screen "IGG Digital Inputs" 1280x800, template "Template"
   on GenerateScreen: "TitleUpdater"()
   Button "HmiScreenItemData_1" at 1,1 size 150x43; TextOn 'Back'; TextOff 'Commissioning'
      on Release: ActivateScreen("Commissioning Main Page", 0)
   AlarmView "Alarm view_1" at 0,777 size 1280x23
   TextField "Text field_1" at 315,140 size 55x22; Text 'I0.0'
   TextField "Text field_2" at 315,176 size 55x22; Text 'I0.1'
   TextField "Text field_3" at 315,212 size 55x22; Text 'I0.2'
   TextField "Text field_4" at 315,248 size 55x22; Text 'I0.3'
   TextField "Text field_5" at 315,283 size 55x22; Text 'I0.4'
   TextField "Text field_6" at 315,319 size 55x22; Text 'I0.5'
   TextField "Text field_7" at 315,355 size 55x22; Text 'I0.6'
   TextField "Text field_8" at 315,391 size 55x22; Text 'I0.7'
   Circle "Circle_1" at 375,140 size 20x20
      Appearance <- "10_DI_Data_IGG_ESTOP_OK"
   Circle "Circle_2" at 375,176 size 20x20
      Appearance <- "10_DI_Data_E139_READY"
   Circle "Circle_3" at 375,212 size 20x20
      Appearance <- "10_DI_Data_E500A_TRIPPED"
   Circle "Circle_4" at 375,248 size 20x20
      Appearance <- "10_DI_Data_E500B_TRIPPED(1)"
   Circle "Circle_5" at 375,283 size 20x20
      Appearance <- "10_DI_Data_E500A_ENBLD(1)"
   Circle "Circle_6" at 375,319 size 20x20
      Appearance <- "10_DI_Data_E500B_ENBLD(1)"
   Circle "Circle_7" at 375,355 size 20x20
      Appearance <- "10_DI_Data_CV401_OPN"
   Circle "Circle_8" at 375,391 size 20x20
      Appearance <- "10_DI_Data_CV401_CLSD"
   TextField "Text field_9" at 332,108 size 49x26; Text 'I0'
   TextField "Text field_10" at 315,461 size 55x22; Text 'I1.0'
   TextField "Text field_11" at 315,497 size 55x22; Text 'I1.1'
   TextField "Text field_12" at 315,533 size 55x22; Text 'I1.2'
   TextField "Text field_13" at 315,569 size 55x22; Text 'I1.3'
   TextField "Text field_14" at 315,604 size 55x22; Text 'I1.4'
   TextField "Text field_15" at 315,640 size 55x22; Text 'I1.5'
   TextField "Text field_16" at 315,676 size 55x22; Text 'I1.6'
   TextField "Text field_17" at 315,712 size 55x22; Text 'I1.7'
   Circle "Circle_9" at 375,461 size 20x20
      Appearance <- "10_DI_Data_CV321_OPN"
   Circle "Circle_10" at 375,497 size 20x20
      Appearance <- "10_DI_Data_CV321_CLSD"
   Circle "Circle_11" at 375,533 size 20x20
      Appearance <- "10_DI_Data_CV322_OPN"
   Circle "Circle_12" at 375,569 size 20x20
      Appearance <- "10_DI_Data_CV322_CLSD"
   Circle "Circle_13" at 375,604 size 20x20
      Appearance <- "10_DI_Data_CV311_OPN"
   Circle "Circle_14" at 375,640 size 20x20
      Appearance <- "10_DI_Data_CV311_CLSD"
   Circle "Circle_15" at 375,676 size 20x20
      Appearance <- "10_DI_Data_CV312_OPN"
   Circle "Circle_16" at 375,712 size 20x20
      Appearance <- "10_DI_Data_CV312_CLSD"
   TextField "Text field_18" at 332,429 size 49x26; Text 'I1'
   TextField "Text field_19" at 657,141 size 55x22; Text 'I2.0'
   TextField "Text field_20" at 657,177 size 55x22; Text 'I2.1'
   TextField "Text field_21" at 657,213 size 55x22; Text 'I2.2'
   TextField "Text field_22" at 657,249 size 55x22; Text 'I2.3'
   TextField "Text field_23" at 657,284 size 55x22; Text 'I2.4'
   TextField "Text field_24" at 657,320 size 55x22; Text 'I2.5'
   TextField "Text field_25" at 657,356 size 55x22; Text 'I2.6'
   TextField "Text field_26" at 657,392 size 55x22; Text 'I2.7'
   Circle "Circle_17" at 717,141 size 20x20
      Appearance <- "10_DI_Data_BC_PLC_PWR_OK"
   Circle "Circle_18" at 717,177 size 20x20
      Appearance <- "10_DI_Data_IGG_VNT_PWR_OK"
   Circle "Circle_19" at 717,213 size 20x20
      Appearance <- "10_DI_Data_MCC_VNT_PWR_OK"
   Circle "Circle_20" at 717,249 size 20x20
      Appearance <- "10_DI_Data_7T1_PWR_OK"
   Circle "Circle_21" at 717,284 size 20x20
      Appearance <- "10_DI_Data_7T2_PWR_OK"
   Circle "Circle_22" at 717,320 size 20x20
      Appearance <- "10_DI_Data_7T3_PWR_OK"
   Circle "Circle_23" at 717,356 size 20x20
      Appearance <- "10_DI_Data_MAINTD_24VDC_PWR_OK"
   Circle "Circle_24" at 717,392 size 20x20
      Appearance <- "10_DI_Data_SFTY_SYS_IL"
   TextField "Text field_27" at 674,109 size 49x26; Text 'I2'
   TextField "Text field_37" at 315,66 size 254x26; Text 'IGG System PLC (Rack 1)'
   TextField "Text field_28" at 657,459 size 55x22; Text 'I3.0'
   TextField "Text field_29" at 657,495 size 55x22; Text 'I3.1'
   TextField "Text field_30" at 657,531 size 55x22; Text 'I3.2'
   TextField "Text field_31" at 657,567 size 55x22; Text 'I3.3'
   TextField "Text field_32" at 657,602 size 55x22; Text 'I3.4'
   TextField "Text field_33" at 657,638 size 55x22; Text 'I3.5'
   TextField "Text field_34" at 657,674 size 55x22; Text 'I3.6'
   TextField "Text field_35" at 657,710 size 55x22; Text 'I3.7'
   Circle "Circle_25" at 717,459 size 20x20
      Appearance <- "10_DI_Data_CV432_OPN"
   Circle "Circle_26" at 717,495 size 20x20
      Appearance <- "10_DI_Data_CV432_CLSD"
   Circle "Circle_27" at 717,531 size 20x20
      Appearance <- "10_DI_Data_CV431_OPN"
   Circle "Circle_28" at 717,567 size 20x20
      Appearance <- "10_DI_Data_CV431_CLSD"
   Circle "Circle_29" at 717,602 size 20x20
      Appearance <- "10_DI_Data_E139_RUNNING(1)"
   Circle "Circle_30" at 717,638 size 20x20
      Appearance <- "10_DI_Data_E139_VSD_FLT"
   Circle "Circle_31" at 717,674 size 20x20
      Appearance <- "10_DI_Data_MCCP_5PG1_OK"
   Circle "Circle_32" at 717,710 size 20x20
      Appearance <- "10_DI_Data_R1_SPR_DI_3_7"
   TextField "Text field_36" at 674,427 size 49x26; Text 'I3'
   TextField "Text field_75" at 408,140 size 200x22; Text 'IGG E-Stop Healthy'
   TextField "Text field_76" at 408,175 size 200x22; Text 'CA Blower Ready E139'
   TextField "Text field_77" at 408,211 size 200x22; Text 'Fuel Pump 1 Tripped E500A'
   TextField "Text field_78" at 408,247 size 200x22; Text 'Fuel Pump 2 Tripped E500B'
   TextField "Text field_79" at 408,283 size 200x22; Text 'Fuel Pump 1 Enabled E500A'
   TextField "Text field_80" at 408,319 size 200x22; Text 'Fuel Pump 2 Enabled E500B'
   TextField "Text field_81" at 408,355 size 200x22; Text 'IG Supply Valve Open CV401'
   TextField "Text field_82" at 408,391 size 200x22; Text 'IG Supply Valve Closed CV401'
   TextField "Text field_83" at 408,460 size 200x22; Text 'DTB Valve Open CV321'
   TextField "Text field_84" at 408,496 size 200x22; Text 'DTB Valve Closed CV321'
   TextField "Text field_85" at 408,532 size 200x22; Text 'CSW Drain Valve Open CV322'
   TextField "Text field_86" at 408,568 size 200x22; Text 'CSW Drain Valve Closed CV322'
   TextField "Text field_87" at 408,604 size 200x22; Text 'CSW Valve Open CV311'
   TextField "Text field_88" at 408,640 size 200x22; Text 'CSW Valve Closed CV311'
   TextField "Text field_89" at 408,676 size 200x22; Text 'Flue Gas S CSW Valve Open CV312'
   TextField "Text field_90" at 408,712 size 200x22; Text 'Flue Gas S CSW Valve Closed CV312'
   TextField "Text field_91" at 748,139 size 200x22; Text 'BC PLC Power Healthy'
   TextField "Text field_92" at 748,175 size 200x22; Text 'IGG Vent Power Healthy'
   TextField "Text field_93" at 748,211 size 200x22; Text 'MCC Vent Power Healthy'
   TextField "Text field_94" at 748,247 size 200x22; Text '7T1 Power Healthy'
   TextField "Text field_95" at 748,283 size 200x22; Text '7T2 Power Healthy'
   TextField "Text field_96" at 748,319 size 200x22; Text '7T3 Power Healthy'
   TextField "Text field_97" at 748,355 size 200x22; Text 'Maintained 24V Power'
   TextField "Text field_98" at 748,392 size 200x22; Text 'Safety System Interlock'
   TextField "Text field_99" at 749,458 size 200x22; Text 'CB IG Supply Valve Open CV432'
   TextField "Text field_100" at 749,494 size 200x22; Text 'CB IG Supply Valve Closed CV432'
   TextField "Text field_101" at 749,530 size 200x22; Text 'BWTS IG Supply Open CV431'
   TextField "Text field_102" at 749,566 size 200x22; Text 'BWTS IG Supply Closed CV431'
   TextField "Text field_103" at 749,602 size 200x22; Text 'CA Blower Running E139'
   TextField "Text field_104" at 749,638 size 200x22; Text 'VSD Fault'
   TextField "Text field_105" at 749,674 size 200x22; Text 'Correct Phase Rotation'
   TextField "Text field_106" at 749,711 size 200x22; Text 'Spare Input'
   Group "Group" at 750,42 size 373x50
   Button "HmiScreenItemData_8" at 764,46 size 355x40; TextOn 'Back'; TextOff 'Text'
   TextField "Screen title" at 750,42 size 373x50; Text 'Screen title'

screen "BC Digital Outputs" 1280x800, template "Template"
   on GenerateScreen: "TitleUpdater"()
   Button "HmiScreenItemData_1" at 1,1 size 150x43; TextOn 'Back'; TextOff 'Commissioning'
      on Release: ActivateScreen("Commissioning Main Page", 0)
   AlarmView "Alarm view_1" at 0,777 size 1280x23
   TextField "Text field_37" at 319,170 size 287x26; Text 'Burner Control PLC (Rack 2)'
   TextField "Text field_38" at 384,239 size 55x22; Text 'Q0.0'
   TextField "Text field_39" at 384,290 size 55x22; Text 'Q0.1'
   TextField "Text field_40" at 384,342 size 55x22; Text 'Q0.2'
   TextField "Text field_41" at 384,394 size 55x22; Text 'Q0.3'
   TextField "Text field_42" at 384,446 size 55x22; Text 'Q0.4'
   TextField "Text field_43" at 384,498 size 55x22; Text 'Q0.5'
   TextField "Text field_44" at 384,550 size 55x22; Text 'Q0.6'
   TextField "Text field_45" at 384,602 size 55x22; Text 'Q0.7'
   Circle "Circle_33" at 443,239 size 20x20
      Appearance <- "14_DQ_Data_200CV127ControlOut"
   Circle "Circle_34" at 443,290 size 20x20
      Appearance <- "14_DQ_Data_200CV124ControlOut"
   Circle "Circle_35" at 443,342 size 20x20
      Appearance <- "14_DQ_Data_200CV215ControlOut"
   Circle "Circle_36" at 443,394 size 20x20
      Appearance <- "14_DQ_Data_200CV216ControlOut"
   Circle "Circle_37" at 443,446 size 20x20
      Appearance <- "14_DQ_Data_200CV114ControlOut"
   Circle "Circle_38" at 443,498 size 20x20
      Appearance <- "14_DQ_Data_200CV206ControlOut"
   Circle "Circle_39" at 443,550 size 20x20
      Appearance <- "14_DQ_Data_200CV207ControlOut"
   Circle "Circle_40" at 443,602 size 20x20
      Appearance <- "14_DQ_Data_E131ControlOut"
   TextField "Text field_46" at 398,206 size 49x26; Text 'Q0'
   TextField "Text field_47" at 703,239 size 55x22; Text 'Q1.0'
   TextField "Text field_48" at 703,290 size 55x22; Text 'Q1.1'
   TextField "Text field_49" at 703,342 size 55x22; Text 'Q1.2'
   TextField "Text field_50" at 703,394 size 55x22; Text 'Q1.3'
   TextField "Text field_51" at 703,446 size 55x22; Text 'Q1.4'
   TextField "Text field_52" at 703,498 size 55x22; Text 'Q1.5'
   TextField "Text field_53" at 703,550 size 55x22; Text 'Q1.6'
   TextField "Text field_54" at 703,602 size 55x22; Text 'Q1.7'
   Circle "Circle_41" at 763,239 size 20x20
      Appearance <- "51_SLAVE_STATUS_P301_ENBLD"
   Circle "Circle_42" at 763,290 size 20x20
      Appearance <- "14_DQ_Data_X001ControlOut"
   Circle "Circle_43" at 763,341 size 20x20
      Appearance <- "14_DQ_Data_R2_SPR_DQ_1_2"
   Circle "Circle_44" at 763,394 size 20x20
      Appearance <- "14_DQ_Data_R2_SPR_DQ_1_3"
   Circle "Circle_45" at 763,446 size 20x20
      Appearance <- "14_DQ_Data_R2_SPR_DQ_1_4"
   Circle "Circle_46" at 763,500 size 20x20
      Appearance <- "14_DQ_Data_R2_SPR_DQ_1_5"
   Circle "Circle_47" at 763,551 size 20x20
      Appearance <- "14_DQ_Data_R2_SPR_DQ_1_6"
   Circle "Circle_48" at 763,602 size 20x20
      Appearance <- "14_DQ_Data_P305ControlOut"
   TextField "Text field_55" at 716,206 size 49x26; Text 'Q1'
   Button "Button_1" at 321,231 size 60x35; TextOff 'Override'
      on Press: InvertBit("80_From_HMI_MAN_DQ_0_0(1)")
      Visibility <- "82_To_HMI_CRNT_MODE_IGG"
   Button "Button_2" at 321,283 size 60x35; TextOff 'Override'
      on Press: InvertBit("80_From_HMI_MAN_DQ_0_1(1)")
      Visibility <- "82_To_HMI_CRNT_MODE_IGG"
   Button "Button_3" at 321,335 size 60x35; TextOff 'Override'
      on Press: InvertBit("80_From_HMI_MAN_DQ_0_2(1)")
      Visibility <- "82_To_HMI_CRNT_MODE_IGG"
   Button "Button_4" at 321,387 size 60x35; TextOff 'Override'
      on Press: InvertBit("80_From_HMI_MAN_DQ_0_3(1)")
      Visibility <- "82_To_HMI_CRNT_MODE_IGG"
   Button "Button_5" at 321,439 size 60x35; TextOff 'Override'
      on Press: InvertBit("80_From_HMI_MAN_DQ_0_4(1)")
      Visibility <- "82_To_HMI_CRNT_MODE_IGG"
   Button "Button_6" at 321,491 size 60x35; TextOff 'Override'
      on Press: InvertBit("80_From_HMI_MAN_DQ_0_5(1)")
      Visibility <- "82_To_HMI_CRNT_MODE_IGG"
   Button "Button_7" at 321,543 size 60x35; TextOff 'Override'
      on Press: InvertBit("80_From_HMI_MAN_DQ_0_6(1)")
      Visibility <- "82_To_HMI_CRNT_MODE_IGG"
   Button "Button_8" at 639,283 size 60x35; TextOff 'Override'
      on Press: InvertBit("80_From_HMI_MAN_DQ_1_1(1)")
      Visibility <- "82_To_HMI_CRNT_MODE_IGG"
   Button "Button_13" at 321,596 size 60x35; TextOff 'Override'
      on Press: InvertBit("80_From_HMI_MAN_DQ_0_7")
      Visibility <- "82_To_HMI_CRNT_MODE_IGG"
   TextField "Text field_72" at 465,239 size 170x22; Text 'Test Pressure Valve CV127'
   TextField "Text field_73" at 465,290 size 170x22; Text 'Pilot B Ign Valve CV124'
   TextField "Text field_75" at 465,342 size 170x22; Text 'Pilot B Fuel Valve 1 CV215'
   TextField "Text field_76" at 465,394 size 170x22; Text 'Pilot B Fuel Valve 2 CV215'
   TextField "Text field_77" at 465,446 size 170x22; Text 'Main B Atom Air Vlv CV114'
   TextField "Text field_78" at 465,498 size 170x22; Text 'Main B Fuel Valve 1 CV205'
   TextField "Text field_79" at 465,550 size 170x22; Text 'Main B Fuel Valve 2 CV206'
   TextField "Text field_80" at 465,602 size 170x22; Text 'IA Comp E131'
   TextField "Text field_81" at 792,238 size 170x22; Text 'CSW Pump P301'
   TextField "Text field_82" at 792,290 size 170x22; Text 'Ignitor X001'
   TextField "Text field_86" at 792,342 size 170x22; Text 'Spare Output'
   TextField "Text field_87" at 792,394 size 170x22; Text 'Spare Output'
   TextField "Text field_88" at 792,446 size 170x22; Text 'Spare Output'
   TextField "Text field_89" at 792,498 size 170x22; Text 'Spare Output'
   TextField "Text field_90" at 792,550 size 170x22; Text 'Spare Output'
   TextField "Text field_91" at 792,602 size 170x22; Text 'Fresh Water Pump'
   Button "Button_26" at 639,231 size 60x35; TextOff 'Override'
      on Press: InvertBit("80_From_HMI_MAN_DQ_1_0")
      Visibility <- "82_To_HMI_CRNT_MODE_IGG"
   Button "Button_27" at 639,335 size 60x35; TextOff 'Override'
      on Press: InvertBit("80_From_HMI_MAN_DQ_1_2(1)")
      Visibility <- "82_To_HMI_CRNT_MODE_IGG"
   Button "Button_28" at 639,439 size 60x35; TextOff 'Override'
      on Press: InvertBit("80_From_HMI_MAN_DQ_1_4(1)")
      Visibility <- "82_To_HMI_CRNT_MODE_IGG"
   Button "Button_29" at 639,387 size 60x35; TextOff 'Override'
      on Press: InvertBit("80_From_HMI_MAN_DQ_1_3(1)")
      Visibility <- "82_To_HMI_CRNT_MODE_IGG"
   Button "Button_30" at 639,491 size 60x35; TextOff 'Override'
      on Press: InvertBit("80_From_HMI_MAN_DQ_1_5(1)")
      Visibility <- "82_To_HMI_CRNT_MODE_IGG"
   Button "Button_31" at 639,543 size 60x35; TextOff 'Override'
      on Press: InvertBit("80_From_HMI_MAN_DQ_1_6")
      Visibility <- "82_To_HMI_CRNT_MODE_IGG"
   Button "Button_32" at 639,596 size 60x35; TextOff 'Override'
      on Press: InvertBit("80_From_HMI_MAN_DQ_1_7(1)")
      Visibility <- "82_To_HMI_CRNT_MODE_IGG"
   Group "Group" at 455,41 size 373x50
   Button "HmiScreenItemData_8" at 469,45 size 355x40; TextOn 'Back'; TextOff 'Text'
   TextField "Screen title" at 455,41 size 373x50; Text 'Screen title'

screen "BC Analogue Inputs" 1280x800, template "Template"
   on GenerateScreen: "TitleUpdater"()
   Button "HmiScreenItemData_1" at 1,1 size 150x43; TextOn 'Back'; TextOff 'Commissioning'
      on Release: ActivateScreen("Commissioning Main Page", 0)
   Button "Button_1" at 34,732 size 100x35; TextOn 'BWTS Digital Inputs'; TextOff 'Back'
      on Click: ActivateScreen("IGG Analogue Inputs", 0)
   TextField "Text field_39" at 34,688 size 171x62; Text 'To IGG Analogue Inputs'
   AlarmView "Alarm view_1" at 0,777 size 1280x23
   Group "Group_1" at 455,41 size 373x50
   TextField "Text field_26" at 607,234 size 64x20; Text 'Reading'
   TextField "Text field_27" at 680,234 size 68x20; Text 'Low Low'
   TextField "Text field_28" at 761,234 size 37x20; Text 'Low'
   TextField "Text field_29" at 829,234 size 37x20; Text 'High'
   TextField "Text field_30" at 879,234 size 74x20; Text 'High High'
   TextField "Text field_31" at 755,211 size 76x20; Text 'Setpoints'
   TextField "Text field_42" at 450,234 size 89x20; Text 'Description'
   TextField "Text field_44" at 340,234 size 37x20; Text 'AI'
   TextField "Text field_53" at 335,202 size 364x26; Text 'Burner Control System PLC (Rack 2)'
   TextField "Text field_35" at 381,576 size 220x22; Text 'E-700 - Inert Gas Soot Content'
   IOField "I/O field_61" at 608,576 size 70x22; FormatPattern 999.99; Unit  %
      ProcessValue <- "12_AI_Data_E700SootContentIn"
   IOField "I/O field_62" at 682,576 size 60x22; FormatPattern 9.9
   TextField "Text field_36" at 328,576 size 50x22; Text 'IW110'
   IOField "I/O field_64" at 750,576 size 60x22; Authorization "Parameter Change"; FormatPattern 99.9
      ProcessValue <- "84_Setpoints_TX700_Low"
   IOField "I/O field_65" at 818,576 size 60x22; Authorization "Parameter Change"; FormatPattern 99.9
      ProcessValue <- "84_Setpoints_TX700_High"
   IOField "I/O field_63" at 886,576 size 60x22; FormatPattern 9.9
   TextField "Text field_1" at 381,536 size 220x22; Text 'E-600 CB - Oxygen Analyser Content'
   IOField "I/O field_2" at 750,536 size 60x22; Authorization "Parameter Change"; FormatPattern 9.99
      ProcessValue <- "84_Setpoints_E600_CB_Low"
   TextField "Text field_2" at 328,536 size 50x22; Text 'IW108'
   IOField "I/O field_8" at 818,536 size 60x22; Authorization "Parameter Change"; FormatPattern 9.99
      ProcessValue <- "84_Setpoints_E600_CB_High"
   IOField "I/O field_1" at 682,536 size 60x22; Authorization "Parameter Change"; FormatPattern 9.99
      ProcessValue <- "84_Setpoints_E600_CB_LowLow"
   IOField "I/O field_9" at 886,536 size 60x22; Authorization "Parameter Change"; FormatPattern 9.99
      ProcessValue <- "84_Setpoints_E600_CB_HighHigh"
   TextField "Text field_33" at 381,496 size 220x22; Text 'E-600 BWTS - Oxygen Analyser Content'
   IOField "I/O field_56" at 608,496 size 70x22; FormatPattern 99.99; Unit  %
      ProcessValue <- "12_AI_Data_E600O2ContentIn"
   IOField "I/O field_58" at 750,496 size 60x22; Authorization "Parameter Change"; FormatPattern 9.99
      ProcessValue <- "84_Setpoints_E600_BWT_Low"
   TextField "Text field_34" at 328,496 size 50x22; Text 'IW108'
   IOField "I/O field_59" at 818,496 size 60x22; Authorization "Parameter Change"; FormatPattern 9.99
      ProcessValue <- "84_Setpoints_E600_BWT_High"
   IOField "I/O field_10" at 886,496 size 60x22; Authorization "Parameter Change"; FormatPattern 9.99
      ProcessValue <- "84_Setpoints_E600_BWT_HighHigh"
   IOField "I/O field_11" at 682,496 size 60x22; Authorization "Parameter Change"; FormatPattern 9.99
      ProcessValue <- "84_Setpoints_E600_BWT_LowLow"
   TextField "Text field_25" at 381,456 size 220x22; Text 'TIT-202 - Inlet Fuel Temperature'
   IOField "I/O field_51" at 608,456 size 70x22; FormatPattern s999.9; Unit  °C
      ProcessValue <- "12_AI_Data_TIT202In_SCALED"
   TextField "Text field_32" at 328,456 size 50x22; Text 'IW106'
   IOField "I/O field_52" at 682,456 size 60x22; Authorization "Parameter Change"; FormatPattern s999.9
      ProcessValue <- "84_Setpoints_TIT202_LowLow"
   IOField "I/O field_53" at 750,456 size 60x22; Authorization "Parameter Change"; FormatPattern s999.9
      ProcessValue <- "84_Setpoints_TIT202_Low"
   IOField "I/O field_54" at 818,456 size 60x22; Authorization "Parameter Change"; FormatPattern s999.9
      ProcessValue <- "84_Setpoints_TIT202_High"
   IOField "I/O field_55" at 886,456 size 60x22; Authorization "Parameter Change"; FormatPattern s999.9
      ProcessValue <- "84_Setpoints_TIT202_HighHigh"
   TextField "Text field_73" at 381,417 size 220x22; Text 'PIT-204 - IGG Inlet Fuel Pressure'
   IOField "I/O field_146" at 608,417 size 70x22; FormatPattern 99.9; Unit  Bar
      ProcessValue <- "12_AI_Data_PIT204In_SCALED"
   TextField "Text field_74" at 328,417 size 50x22; Text 'IW104'
   IOField "I/O field_147" at 682,417 size 60x22; Authorization "Parameter Change"; FormatPattern 99.9
      ProcessValue <- "84_Setpoints_PIT204_LowLow(2)"
   IOField "I/O field_148" at 750,417 size 60x22; Authorization "Parameter Change"; FormatPattern 99.9
      ProcessValue <- "84_Setpoints_PIT204_Low(2)"
   IOField "I/O field_149" at 818,417 size 60x22; Authorization "Parameter Change"; FormatPattern 99.9
      ProcessValue <- "84_Setpoints_PIT204_High(2)"
   IOField "I/O field_150" at 886,417 size 60x22; Authorization "Parameter Change"; FormatPattern 99.9
      ProcessValue <- "84_Setpoints_PIT204_HighHigh(2)"
   TextField "Text field_71" at 381,378 size 220x22; Text 'PIT-112 - Inlet IA Compressor Pressure'
   TextField "Text field_72" at 328,378 size 50x22; Text 'IW102'
   IOField "I/O field_3" at 608,378 size 70x22; FormatPattern 99.9; Unit  Bar
      ProcessValue <- "12_AI_Data_PIT112In_SCALED"
   IOField "I/O field_4" at 682,378 size 60x22; Authorization "Parameter Change"; FormatPattern 99.9
      ProcessValue <- "84_Setpoints_PIT112_LowLow"
   IOField "I/O field_5" at 750,378 size 60x22; Authorization "Parameter Change"; FormatPattern 99.9
      ProcessValue <- "84_Setpoints_PIT112_Low"
   IOField "I/O field_6" at 818,378 size 60x22; Authorization "Parameter Change"; FormatPattern 99.9
      ProcessValue <- "84_Setpoints_PIT112_High"
   IOField "I/O field_7" at 886,378 size 60x22; Authorization "Parameter Change"; FormatPattern 99.9
      ProcessValue <- "84_Setpoints_PIT112_HighHigh"
   TextField "Text field_69" at 381,338 size 220x22; Text 'PIT-113 - Main Atom. Air Pressure'
   IOField "I/O field_136" at 608,338 size 70x22; FormatPattern 99.9; Unit  Bar
      ProcessValue <- "12_AI_Data_PIT113In_SCALED"
   TextField "Text field_70" at 328,338 size 50x22; Text 'IW100'
   IOField "I/O field_137" at 682,338 size 60x22; Authorization "Parameter Change"; FormatPattern 99.9
      ProcessValue <- "84_Setpoints_PIT113_LowLow"
   IOField "I/O field_138" at 750,338 size 60x22; Authorization "Parameter Change"; FormatPattern 99.9
      ProcessValue <- "84_Setpoints_PIT113_Low"
   IOField "I/O field_139" at 818,338 size 60x22; Authorization "Parameter Change"; FormatPattern 99.9
      ProcessValue <- "84_Setpoints_PIT113_High"
   IOField "I/O field_140" at 886,338 size 60x22; Authorization "Parameter Change"; FormatPattern 99.9
      ProcessValue <- "84_Setpoints_PIT113_HighHigh"
   TextField "Text field_67" at 381,299 size 220x22; Text 'FD-001 - Flame Signal'
   IOField "I/O field_131" at 608,299 size 70x22; FormatPattern 999.9; Unit  %
      ProcessValue <- "12_AI_Data_FD001FlameSignalIn"
   IOField "I/O field_134" at 818,299 size 60x22; FormatPattern s99.9
   IOField "I/O field_135" at 886,299 size 60x22; FormatPattern s99.9
   TextField "Text field_68" at 328,299 size 50x22; Text 'IW98'
   IOField "I/O field_132" at 682,299 size 60x22; Authorization "Parameter Change"; FormatPattern 999.9
      ProcessValue <- "84_Setpoints_FD001_LowLow"
   IOField "I/O field_133" at 750,299 size 60x22; Authorization "Parameter Change"; FormatPattern 999.9
      ProcessValue <- "84_Setpoints_FD001_Low"
   TextField "Text field_65" at 381,260 size 220x22; Text 'PIT-205 - IGG Main Fuel Pressure'
   IOField "I/O field_126" at 608,260 size 70x22; FormatPattern 99.9; Unit  Bar
      ProcessValue <- "12_AI_Data_PIT205In_SCALED"
   TextField "Text field_66" at 328,260 size 50x22; Text 'IW96'
   IOField "I/O field_127" at 682,260 size 60x22; Authorization "Parameter Change"; FormatPattern 99.9
      ProcessValue <- "84_Setpoints_PIT205_LowLow"
   IOField "I/O field_128" at 750,260 size 60x22; Authorization "Parameter Change"; FormatPattern 99.9
      ProcessValue <- "84_Setpoints_PIT205_Low"
   IOField "I/O field_129" at 818,260 size 60x22; Authorization "Parameter Change"; FormatPattern 99.9
      ProcessValue <- "84_Setpoints_PIT205_High"
   IOField "I/O field_130" at 886,260 size 60x22; Authorization "Parameter Change"; FormatPattern 99.9
      ProcessValue <- "84_Setpoints_PIT205_HighHigh"
   Button "HmiScreenItemData_8" at 469,45 size 355x40; TextOn 'Back'; TextOff 'Text'
   TextField "Screen title" at 455,41 size 373x50; Text 'Screen title'

screen "IGG Analogue Outputs" 1280x800, template "Template"
   on GenerateScreen: "TitleUpdater"()
   Button "HmiScreenItemData_1" at 1,1 size 150x43; TextOn 'Back'; TextOff 'Commissioning'
      on Release: ActivateScreen("Commissioning Main Page", 0)
   Button "Button_15" at 34,732 size 100x35; TextOn 'BWTS Digital Inputs'; TextOff 'Back'
      on Click: ActivateScreen("BC Analogue Inputs", 0)
   AlarmView "Alarm view_1" at 0,777 size 1280x23
   TextField "Text field_82" at 481,361 size 220x22; Text 'Vent Valve Position Control'
   TextField "Text field_90" at 750,332 size 64x20; Text 'Reading'
   IOField "I/O field_2" at 749,363 size 70x22; FormatPattern 9999; Unit %
      ProcessValue <- "16_AQ_Data_CV403_CNTRL"
   TextField "Text field_6" at 428,361 size 53x22; Text 'QW98'
   TextField "Text field_7" at 480,438 size 220x22; Text 'Spare'
   TextField "Text field_41" at 553,332 size 89x20; Text 'Description'
   TextField "Text field_43" at 437,332 size 37x20; Text 'AO'
   TextField "Text field_52" at 437,299 size 333x26; Text 'IGG Control System PLC (Rack 1)'
   TextField "Text field_25" at 480,399 size 220x22; Text 'CA Blower Speed Control'
   IOField "I/O field_51" at 749,398 size 70x22; FormatPattern 9999; Unit RPM
      ProcessValue <- "16_AQ_Data_E139_SPEED"
   TextField "Text field_32" at 427,399 size 53x22; Text 'QW100'
   Button "Button_24" at 716,359 size 29x26; TextOff '+'
      Visibility <- "82_To_HMI_CRNT_MODE_IGG"
      on Press: function_b14e0dd5("80_From_HMI_MAN_AQ_INC_98(1)", 0)
   Button "Button_25" at 824,359 size 29x26; TextOff '-'
      Visibility <- "82_To_HMI_CRNT_MODE_IGG"
      on Press: function_b14e0dd5("80_From_HMI_MAN_AQ_DEC_98(1)", 0)
   Button "Button_1" at 717,397 size 29x26; TextOff '+'
      Visibility <- "82_To_HMI_CRNT_MODE_IGG"
      on Press: function_b14e0dd5("80_From_HMI_MAN_AQ_INC_100", 0)
   Button "Button_2" at 825,397 size 29x26; TextOff '-'
      Visibility <- "82_To_HMI_CRNT_MODE_IGG"
      on Press: function_b14e0dd5("80_From_HMI_MAN_AQ_DEC_100", 0)
   Button "Button_3" at 715,434 size 29x26; TextOff '+'
      on Click: SetBit("80_From_HMI_MAN_AQ_INC_102(1)")
      Visibility <- "82_To_HMI_CRNT_MODE_IGG"
   Button "Button_4" at 823,434 size 29x26; TextOff '-'
      on Click: SetBit("80_From_HMI_MAN_AQ_DEC_102(1)")
      Visibility <- "82_To_HMI_CRNT_MODE_IGG"
   Button "Button_5" at 716,475 size 29x26; TextOff '+'
      on Click: SetBit("80_From_HMI_MAN_AQ_INC_104")
      Visibility <- "82_To_HMI_CRNT_MODE_IGG"
   Button "Button_6" at 824,475 size 29x26; TextOff '-'
      on Click: SetBit("80_From_HMI_MAN_AQ_DEC_104")
      Visibility <- "82_To_HMI_CRNT_MODE_IGG"
   IOField "I/O field_1" at 749,438 size 70x22; FormatPattern 9.9; Unit  
      ProcessValue <- "16_AQ_Data_R1_SPR_AQ_102"
   IOField "I/O field_3" at 750,478 size 70x22; FormatPattern 9.9; Unit  
      ProcessValue <- "16_AQ_Data_R1_SPR_AQ_104"
   TextField "Text field_1" at 480,478 size 220x22; Text 'Spare'
   TextField "Text field_2" at 428,438 size 53x22; Text 'QW102'
   TextField "Text field_3" at 427,478 size 53x22; Text 'QW104'
   Group "Group" at 455,41 size 373x50
   Button "HmiScreenItemData_8" at 469,45 size 355x40; TextOn 'Back'; TextOff 'Text'
   TextField "Screen title" at 455,41 size 373x50; Text 'Screen title'

screen "IGG Target Setpoints" 1280x800, template "Template"
   on GenerateScreen: "TitleUpdater"()
   Button "HmiScreenItemData_1" at 1,1 size 150x43; TextOn 'Back'; TextOff 'Commissioning'
      on Release: ActivateScreen("Commissioning Main Page", 0)
   AlarmView "Alarm view_1" at 0,777 size 1280x23
   TextField "Text field_25" at 394,430 size 407x22; Text 'PIT-113: IGG Main Atom Air Pressure Target'
   TextField "Text field_29" at 814,210 size 68x20; Text 'Setpoint'
   TextField "Text field_33" at 393,468 size 408x22; Text 'PIT-205: IGG Main Fuel Pressure Target'
   IOField "I/O field_58" at 816,468 size 60x22; Authorization "Parameter Change"; FormatPattern 999.99
      ProcessValue <- "84_Setpoints_PIT205_Target(1)"
   TextField "Text field_35" at 394,552 size 406x22; Text 'E-600: O2 Cargo Blanketing Target'
   TextField "Text field_65" at 394,236 size 411x22; Text 'PIT-402: IG Outlet Pressure Pilot Target'
   TextField "Text field_67" at 394,274 size 410x22; Text 'PIT-402: IG Outlet Pressure Main Target'
   TextField "Text field_69" at 395,313 size 407x22; Text 'PIT-402: IG Outlet Pressure Post Target Start'
   TextField "Text field_71" at 395,352 size 406x22; Text 'PIT-402: IG Outlet Pressure Post Target Maximum'
   TextField "Text field_73" at 395,391 size 407x22; Text 'FD-001: Igniter Target'
   TextField "Text field_42" at 394,210 size 89x20; Text 'Description'
   IOField "I/O field_128" at 816,236 size 60x22; Authorization "Parameter Change"; FormatPattern 999.9
      ProcessValue <- "84_Setpoints_PIT402_Pilot_Target(1)"
   IOField "I/O field_133" at 816,274 size 60x22; Authorization "Parameter Change"; FormatPattern 999.9
      ProcessValue <- "84_Setpoints_PIT402_Main_Target(1)"
   IOField "I/O field_138" at 816,313 size 60x22; Authorization "Parameter Change"; FormatPattern 999.9
      ProcessValue <- "84_Setpoints_PIT402_Post_Target_Start"
   IOField "I/O field_53" at 816,430 size 60x22; Authorization "Parameter Change"; FormatPattern 999.9
      ProcessValue <- "84_Setpoints_PIT113_Pilot_Target(1)"
   IOField "I/O field_148" at 816,391 size 60x22; Authorization "Parameter Change"; FormatPattern 999.9
      ProcessValue <- "84_Setpoints_FD001_Min"
   IOField "I/O field_64" at 816,552 size 60x22; Authorization "Parameter Change"; FormatPattern 99.9
      ProcessValue <- "84_Setpoints_E600_CB_Target"
   TextField "Text field_53" at 393,184 size 213x26; Text 'IGG Target Setpoints'
   IOField "I/O field_5" at 815,352 size 60x22; Authorization "Parameter Change"; FormatPattern 999.9
      ProcessValue <- "84_Setpoints_PIT401_Post_Target_Max"
   TextField "Text field_1" at 394,510 size 406x22; Text 'E-600: O2 Ballast Water Treatment Target'
   IOField "I/O field_2" at 816,510 size 60x22; Authorization "Parameter Change"; FormatPattern 9.99
      ProcessValue <- "84_Setpoints_E600_BWT_Target"
   TextField "Text field_2" at 394,595 size 406x22; Text 'PIT-402 Target Ramp Time (s)'
   IOField "I/O field_1" at 816,595 size 60x22; Authorization "Parameter Change"; FormatPattern 999
      ProcessValue <- "86_Times_PIT402_Ramp_Seconds"
   Group "Group" at 455,41 size 373x50
   Button "HmiScreenItemData_8" at 469,45 size 355x40; TextOn 'Back'; TextOff 'Text'
   TextField "Screen title" at 455,41 size 373x50; Text 'Screen title'

screen "IGG Process Times" 1280x800, template "Template"
   on GenerateScreen: "TitleUpdater"()
   Button "HmiScreenItemData_1" at 1,1 size 150x43; TextOn 'Back'; TextOff 'Commissioning'
      on Release: ActivateScreen("Commissioning Main Page", 0)
   Button "Button_1" at 21,736 size 161x32; TextOff 'IGG Step Times'
      on Activate: ActivateScreen("IGG Max Step Times", 0)
   Button "Button_2" at 1091,736 size 161x32; TextOff 'BC Step Times'
      on Activate: ActivateScreen("BC Max Step Times", 0)
   AlarmView "Alarm view_1" at 0,777 size 1280x23
   TextField "Text field_25" at 458,325 size 286x22; Text 'CV311 Maximum Travel Time'
   TextField "Text field_29" at 758,159 size 65x20; Text 'Time (s)'
   TextField "Text field_33" at 458,353 size 286x22; Text 'CV312 Maximum Travel Time'
   IOField "I/O field_58" at 757,353 size 60x22; Authorization "Parameter Change"; FormatPattern 999
      ProcessValue <- "86_Times_CV312_MAX_TRVL_TIME"
   TextField "Text field_35" at 458,409 size 283x22; Text 'CV322 Maximum Travel Time'
   TextField "Text field_65" at 458,185 size 289x22; Text 'Burner Control Start Command Delay Time'
   TextField "Text field_67" at 458,213 size 288x22; Text 'CV203 Close Command Delay Time'
   TextField "Text field_69" at 458,241 size 287x22; Text 'Post P301 Stopped Delay Time'
   TextField "Text field_71" at 458,269 size 286x22; Text 'Post CV311 Closed Delay Time'
   TextField "Text field_73" at 458,297 size 285x22; Text 'Post CV321 Opened Delay Time'
   TextField "Text field_42" at 458,159 size 89x20; Text 'Description'
   IOField "I/O field_128" at 757,185 size 60x22; Authorization "Parameter Change"; FormatPattern 999
      ProcessValue <- "86_Times_PRE_BC_STRT_CMND_DLY"
   IOField "I/O field_133" at 757,213 size 60x22; Authorization "Parameter Change"; FormatPattern 999
      ProcessValue <- "86_Times_PRE_CV203_CLS_CMND_DLY"
   IOField "I/O field_138" at 757,241 size 60x22; Authorization "Parameter Change"; FormatPattern 999
      ProcessValue <- "86_Times_POST_P301_STOP_DLY"
   IOField "I/O field_148" at 757,298 size 60x22; Authorization "Parameter Change"; FormatPattern 999
      ProcessValue <- "86_Times_POST_CV321_OPN_DLY"
   IOField "I/O field_64" at 757,408 size 60x22; Authorization "Parameter Change"; FormatPattern 999
      ProcessValue <- "86_Times_CV322_MAX_TRVL_TIME"
   TextField "Text field_53" at 457,133 size 190x26; Text 'IGG Process Times'
   IOField "I/O field_5" at 756,270 size 60x22; Authorization "Parameter Change"; FormatPattern 999
      ProcessValue <- "86_Times_POST_CV311_CLS_DLY"
   TextField "Text field_1" at 458,381 size 284x22; Text 'CV321 Maximum Travel Time'
   IOField "I/O field_2" at 757,381 size 60x22; Authorization "Parameter Change"; FormatPattern 999
      ProcessValue <- "86_Times_CV321_MAX_TRVL_TIME"
   TextField "Text field_14" at 458,437 size 283x22; Text 'CV401 Maximum Travel Time'
   IOField "I/O field_12" at 756,439 size 60x22; Authorization "Parameter Change"; FormatPattern 999
      ProcessValue <- "86_Times_CV401_MAX_TRVL_TIME"
   TextField "Text field_15" at 458,465 size 283x22; Text 'CV431 Maximum Travel Time'
   IOField "I/O field_13" at 756,467 size 60x22; Authorization "Parameter Change"; FormatPattern 999
      ProcessValue <- "86_Times_CV431_MAX_TRVL_TIME"
   TextField "Text field_16" at 458,494 size 283x22; Text 'CV432 Maximum Travel Time'
   IOField "I/O field_14" at 756,494 size 60x22; Authorization "Parameter Change"; FormatPattern 999
      ProcessValue <- "86_Times_CV432_MAX_TRVL_TIME"
   IOField "I/O field_15" at 758,326 size 60x22; Authorization "Parameter Change"; FormatPattern 999
      ProcessValue <- "86_Times_CV311_MAX_TRVL_TIME"
   TextField "Text field_44" at 458,524 size 283x22; Text 'FS317 Delayed Fault'
   IOField "I/O field_36" at 756,524 size 60x22; Authorization "Parameter Change"; FormatPattern 999
      ProcessValue <- "86_Times_FS317 delay"
   TextField "Text field_45" at 458,555 size 283x22; Text 'FS320 Delayed Fault'
   IOField "I/O field_37" at 756,555 size 60x22; Authorization "Parameter Change"; FormatPattern 999
      ProcessValue <- "86_Times_FS320 delay"
   TextField "Text field_46" at 458,585 size 283x22; Text 'FS359 Delayed Fault'
   IOField "I/O field_38" at 756,585 size 60x22; Authorization "Parameter Change"; FormatPattern 999
      ProcessValue <- "80_From_HMI_PIT 359 delay"
   TextField "Text field_47" at 458,616 size 283x22; Text 'FS316 Delayed Fault'
   IOField "I/O field_39" at 756,616 size 60x22; Authorization "Parameter Change"; FormatPattern 999
      ProcessValue <- "80_From_HMI_PIT 316 delay"
   TextField "Text field_2" at 458,646 size 283x22; Text 'PIT402 Delayed Fault'
   IOField "I/O field_1" at 756,646 size 60x22; Authorization "Parameter Change"; FormatPattern 999
      ProcessValue <- "86_Times_PIT402 Alarm Delay"
   Group "Group" at 455,41 size 373x50
   Button "HmiScreenItemData_8" at 469,45 size 355x40; TextOn 'Back'; TextOff 'Text'
   TextField "Screen title" at 455,41 size 373x50; Text 'Screen title'

screen "IGG Max Step Times" 1280x800, template "Template"
   on GenerateScreen: "TitleUpdater"()
   Button "HmiScreenItemData_1" at 1,1 size 150x43; TextOn 'Back'; TextOff 'Commissioning'
      on Release: ActivateScreen("Commissioning Main Page", 0)
   TextField "Text field_25" at 101,290 size 286x22; Text 'Step 040'
   TextField "Text field_29" at 401,122 size 77x20; Text 'Time (ms)'
   TextField "Text field_33" at 101,319 size 286x22; Text 'Step 050'
   IOField "I/O field_58" at 400,319 size 60x22; Authorization "Parameter Change"; FormatPattern s9999999999
      ProcessValue <- "86_Times_STEP_MAX_TIME_STP_050(2)"
   TextField "Text field_35" at 101,376 size 283x22; Text 'Step 070'
   TextField "Text field_65" at 101,148 size 289x22; Text 'Step 001'
   TextField "Text field_67" at 101,176 size 288x22; Text 'Step 005'
   TextField "Text field_69" at 101,205 size 287x22; Text 'Step 010'
   TextField "Text field_71" at 101,233 size 286x22; Text 'Step 020'
   TextField "Text field_73" at 101,262 size 285x22; Text 'Step 030'
   TextField "Text field_42" at 101,122 size 89x20; Text 'Description'
   IOField "I/O field_128" at 400,148 size 60x22; Authorization "Parameter Change"; FormatPattern s9999999999
      ProcessValue <- "86_Times_STEP_MAX_TIME_STP_001(2)"
   IOField "I/O field_133" at 400,176 size 60x22; Authorization "Parameter Change"; FormatPattern s9999999999
      ProcessValue <- "86_Times_STEP_MAX_TIME_STP_005(2)"
   IOField "I/O field_138" at 400,205 size 60x22; Authorization "Parameter Change"; FormatPattern s9999999999
      ProcessValue <- "86_Times_STEP_MAX_TIME_STP_010(2)"
   IOField "I/O field_148" at 400,262 size 60x22; Authorization "Parameter Change"; FormatPattern s9999999999
      ProcessValue <- "86_Times_STEP_MAX_TIME_STP_030(2)"
   IOField "I/O field_64" at 400,376 size 60x22; Authorization "Parameter Change"; FormatPattern s9999999999
      ProcessValue <- "86_Times_STEP_MAX_TIME_STP_070(2)"
   TextField "Text field_53" at 100,96 size 259x26; Text 'IGG Maximum Step Times'
   IOField "I/O field_5" at 400,233 size 60x22; Authorization "Parameter Change"; FormatPattern s9999999999
      ProcessValue <- "86_Times_STEP_MAX_TIME_STP_020(2)"
   TextField "Text field_1" at 101,348 size 284x22; Text 'Step 060'
   IOField "I/O field_2" at 400,348 size 60x22; Authorization "Parameter Change"; FormatPattern s9999999999
      ProcessValue <- "86_Times_STEP_MAX_TIME_STP_060(2)"
   TextField "Text field_2" at 479,291 size 271x22; Text 'Step 240'
   TextField "Text field_3" at 768,123 size 77x20; Text 'Time (ms)'
   TextField "Text field_4" at 479,320 size 273x22; Text 'Step 250'
   IOField "I/O field_1" at 767,319 size 60x22; Authorization "Parameter Change"; FormatPattern s9999999999
      ProcessValue <- "86_Times_STEP_MAX_TIME_STP_250(2)"
   TextField "Text field_5" at 479,377 size 270x22; Text 'Step 270'
   TextField "Text field_6" at 479,149 size 272x22; Text 'Step 190'
   TextField "Text field_7" at 479,177 size 272x22; Text 'Step 200'
   TextField "Text field_8" at 479,206 size 271x22; Text 'Step 210'
   TextField "Text field_9" at 479,234 size 270x22; Text 'Step 220'
   TextField "Text field_10" at 479,263 size 270x22; Text 'Step 230'
   TextField "Text field_11" at 479,123 size 89x20; Text 'Description'
   IOField "I/O field_3" at 767,149 size 60x22; Authorization "Parameter Change"; FormatPattern s9999999999
      ProcessValue <- "86_Times_STEP_MAX_TIME_STP_190(2)"
   IOField "I/O field_4" at 767,177 size 60x22; Authorization "Parameter Change"; FormatPattern s9999999999
      ProcessValue <- "86_Times_STEP_MAX_TIME_STP_200(2)"
   IOField "I/O field_6" at 767,205 size 60x22; Authorization "Parameter Change"; FormatPattern s9999999999
      ProcessValue <- "86_Times_STEP_MAX_TIME_STP_210(2)"
   IOField "I/O field_8" at 767,262 size 60x22; Authorization "Parameter Change"; FormatPattern s9999999999
      ProcessValue <- "86_Times_STEP_MAX_TIME_STP_230(2)"
   IOField "I/O field_9" at 767,376 size 60x22; Authorization "Parameter Change"; FormatPattern s9999999999
      ProcessValue <- "86_Times_STEP_MAX_TIME_STP_270(2)"
   IOField "I/O field_10" at 767,234 size 60x22; Authorization "Parameter Change"; FormatPattern s9999999999
      ProcessValue <- "86_Times_STEP_MAX_TIME_STP_220(2)"
   TextField "Text field_13" at 479,348 size 270x22; Text 'Step 260'
   IOField "I/O field_11" at 767,348 size 60x22; Authorization "Parameter Change"; FormatPattern s9999999999
      ProcessValue <- "86_Times_STEP_MAX_TIME_STP_260(2)"
   TextField "Text field_14" at 101,405 size 283x22; Text 'Step 080'
   IOField "I/O field_12" at 400,405 size 60x22; Authorization "Parameter Change"; FormatPattern s9999999999
      ProcessValue <- "86_Times_STEP_MAX_TIME_STP_080(2)"
   TextField "Text field_15" at 101,433 size 283x22; Text 'Step 090'
   IOField "I/O field_13" at 400,433 size 60x22; Authorization "Parameter Change"; FormatPattern s9999999999
      ProcessValue <- "86_Times_STEP_MAX_TIME_STP_090(2)"
   TextField "Text field_16" at 101,462 size 283x22; Text 'Step 100'
   IOField "I/O field_14" at 400,462 size 60x22; Authorization "Parameter Change"; FormatPattern s9999999999
      ProcessValue <- "86_Times_STEP_MAX_TIME_STP_100(2)"
   Button "Button_1" at 21,736 size 161x32; TextOff 'Back'
      on Activate: ActivateScreen("IGG Process Times", 0)
   IOField "I/O field_15" at 400,290 size 60x22; Authorization "Parameter Change"; FormatPattern s9999999999
      ProcessValue <- "86_Times_STEP_MAX_TIME_STP_040(2)"
   TextField "Text field_17" at 479,405 size 270x22; Text 'Step 280'
   IOField "I/O field_16" at 767,405 size 60x22; Authorization "Parameter Change"; FormatPattern s9999999999
      ProcessValue <- "86_Times_STEP_MAX_TIME_STP_280(2)"
   TextField "Text field_18" at 479,434 size 270x22; Text 'Step 290'
   IOField "I/O field_17" at 767,433 size 60x22; Authorization "Parameter Change"; FormatPattern s9999999999
      ProcessValue <- "86_Times_STEP_MAX_TIME_STP_290(2)"
   TextField "Text field_19" at 479,462 size 269x22; Text 'Step 300'
   IOField "I/O field_18" at 767,462 size 60x22; Authorization "Parameter Change"; FormatPattern s9999999999
      ProcessValue <- "86_Times_STEP_MAX_TIME_STP_300(2)"
   TextField "Text field_20" at 479,491 size 269x22; Text 'Step 310'
   IOField "I/O field_19" at 767,490 size 60x22; Authorization "Parameter Change"; FormatPattern s9999999999
      ProcessValue <- "86_Times_STEP_MAX_TIME_STP_310(2)"
   TextField "Text field_21" at 479,519 size 269x22; Text 'Step 320'
   IOField "I/O field_20" at 767,519 size 60x22; Authorization "Parameter Change"; FormatPattern s9999999999
      ProcessValue <- "86_Times_STEP_MAX_TIME_STP_320(2)"
   TextField "Text field_22" at 853,149 size 269x22; Text 'Step 390'
   IOField "I/O field_21" at 1141,149 size 60x22; Authorization "Parameter Change"; FormatPattern s9999999999
      ProcessValue <- "86_Times_STEP_MAX_TIME_STP_390(2)"
   TextField "Text field_23" at 853,122 size 89x20; Text 'Description'
   TextField "Text field_24" at 1140,123 size 77x20; Text 'Time (ms)'
   TextField "Text field_26" at 853,176 size 269x22; Text 'Step 400'
   IOField "I/O field_22" at 1141,176 size 60x22; Authorization "Parameter Change"; FormatPattern s9999999999
      ProcessValue <- "86_Times_STEP_MAX_TIME_STP_400(2)"
   TextField "Text field_27" at 853,204 size 269x22; Text 'Step 410'
   IOField "I/O field_23" at 1141,204 size 60x22; Authorization "Parameter Change"; FormatPattern s9999999999
      ProcessValue <- "86_Times_STEP_MAX_TIME_STP_410(2)"
   TextField "Text field_28" at 853,232 size 269x22; Text 'Step 420'
   IOField "I/O field_24" at 1141,232 size 60x22; Authorization "Parameter Change"; FormatPattern s9999999999
      ProcessValue <- "86_Times_STEP_MAX_TIME_STP_420(2)"
   TextField "Text field_30" at 853,260 size 269x22; Text 'Step 430'
   IOField "I/O field_25" at 1141,260 size 60x22; Authorization "Parameter Change"; FormatPattern s9999999999
      ProcessValue <- "86_Times_STEP_MAX_TIME_STP_430(2)"
   TextField "Text field_31" at 853,288 size 269x22; Text 'Step 440'
   IOField "I/O field_26" at 1141,288 size 60x22; Authorization "Parameter Change"; FormatPattern s9999999999
      ProcessValue <- "86_Times_STEP_MAX_TIME_STP_440(2)"
   TextField "Text field_32" at 853,316 size 269x22; Text 'Step 450'
   IOField "I/O field_27" at 1141,316 size 60x22; Authorization "Parameter Change"; FormatPattern s9999999999
      ProcessValue <- "86_Times_STEP_MAX_TIME_STP_450(2)"
   TextField "Text field_34" at 853,344 size 269x22; Text 'Step 460'
   IOField "I/O field_28" at 1141,344 size 60x22; Authorization "Parameter Change"; FormatPattern s9999999999
      ProcessValue <- "86_Times_STEP_MAX_TIME_STP_460(2)"
   TextField "Text field_36" at 853,372 size 269x22; Text 'Step 470'
   IOField "I/O field_29" at 1141,372 size 60x22; Authorization "Parameter Change"; FormatPattern s9999999999
      ProcessValue <- "86_Times_STEP_MAX_TIME_STP_470(2)"
   TextField "Text field_37" at 853,400 size 269x22; Text 'Step 480'
   IOField "I/O field_30" at 1141,400 size 60x22; Authorization "Parameter Change"; FormatPattern s9999999999
      ProcessValue <- "86_Times_STEP_MAX_TIME_STP_480(2)"
   TextField "Text field_38" at 853,428 size 269x22; Text 'Step 490'
   IOField "I/O field_31" at 1141,428 size 60x22; Authorization "Parameter Change"; FormatPattern s9999999999
      ProcessValue <- "86_Times_STEP_MAX_TIME_STP_490(2)"
   TextField "Text field_39" at 853,456 size 269x22; Text 'Step 500'
   IOField "I/O field_32" at 1141,456 size 60x22; Authorization "Parameter Change"; FormatPattern s9999999999
      ProcessValue <- "86_Times_STEP_MAX_TIME_STP_500(2)"
   IOField "I/O field_7" at 767,291 size 60x22; Authorization "Parameter Change"; FormatPattern s9999999999
      ProcessValue <- "86_Times_STEP_MAX_TIME_STP_240(2)"
   TextField "Text field_43" at 101,490 size 283x22; Text 'Step 110'
   IOField "I/O field_35" at 400,490 size 60x22; Authorization "Parameter Change"; FormatPattern s9999999999
      ProcessValue <- "86_Times_STEP_MAX_TIME_STP_110(2)"
   TextField "Text field_44" at 101,519 size 283x22; Text 'Step 120'
   IOField "I/O field_36" at 400,519 size 60x22; Authorization "Parameter Change"; FormatPattern s9999999999
      ProcessValue <- "86_Times_STEP_MAX_TIME_STP_120(2)"
   TextField "Text field_45" at 479,548 size 269x22; Text 'Step 330'
   IOField "I/O field_37" at 767,547 size 60x22; Authorization "Parameter Change"; FormatPattern s9999999999
      ProcessValue <- "86_Times_STEP_MAX_TIME_STP_330(2)"
   TextField "Text field_47" at 101,548 size 283x22; Text 'Step 130'
   IOField "I/O field_39" at 400,548 size 60x22; Authorization "Parameter Change"; FormatPattern s9999999999
      ProcessValue <- "86_Times_STEP_MAX_TIME_STP_130(2)"
   TextField "Text field_48" at 479,576 size 269x22; Text 'Step 340'
   IOField "I/O field_40" at 767,576 size 60x22; Authorization "Parameter Change"; FormatPattern s9999999999
      ProcessValue <- "86_Times_STEP_MAX_TIME_STP_340(2)"
   TextField "Text field_50" at 101,576 size 283x22; Text 'Step 140'
   IOField "I/O field_42" at 400,576 size 60x22; Authorization "Parameter Change"; FormatPattern s9999999999
      ProcessValue <- "86_Times_STEP_MAX_TIME_STP_140(2)"
   TextField "Text field_51" at 479,605 size 269x22; Text 'Step 350'
   IOField "I/O field_43" at 767,604 size 60x22; Authorization "Parameter Change"; FormatPattern s9999999999
      ProcessValue <- "86_Times_STEP_MAX_TIME_STP_350(2)"
   TextField "Text field_54" at 101,605 size 283x22; Text 'Step 150'
   IOField "I/O field_45" at 400,605 size 60x22; Authorization "Parameter Change"; FormatPattern s9999999999
      ProcessValue <- "86_Times_STEP_MAX_TIME_STP_150(2)"
   TextField "Text field_55" at 479,633 size 269x22; Text 'Step 360'
   IOField "I/O field_46" at 767,633 size 60x22; Authorization "Parameter Change"; FormatPattern s9999999999
      ProcessValue <- "86_Times_STEP_MAX_TIME_STP_360(2)"
   TextField "Text field_57" at 101,633 size 283x22; Text 'Step 160'
   IOField "I/O field_48" at 400,633 size 60x22; Authorization "Parameter Change"; FormatPattern s9999999999
      ProcessValue <- "86_Times_STEP_MAX_TIME_STP_160(2)"
   TextField "Text field_58" at 479,662 size 269x22; Text 'Step 370'
   IOField "I/O field_49" at 767,662 size 60x22; Authorization "Parameter Change"; FormatPattern s9999999999
      ProcessValue <- "86_Times_STEP_MAX_TIME_STP_370(2)"
   TextField "Text field_60" at 101,662 size 283x22; Text 'Step 170'
   IOField "I/O field_51" at 400,662 size 60x22; Authorization "Parameter Change"; FormatPattern s9999999999
      ProcessValue <- "86_Times_STEP_MAX_TIME_STP_170(2)"
   TextField "Text field_61" at 479,691 size 269x22; Text 'Step 380'
   IOField "I/O field_52" at 767,691 size 60x22; Authorization "Parameter Change"; FormatPattern s9999999999
      ProcessValue <- "86_Times_STEP_MAX_TIME_STP_380(2)"
   TextField "Text field_63" at 101,691 size 283x22; Text 'Step 180'
   IOField "I/O field_54" at 400,691 size 60x22; Authorization "Parameter Change"; FormatPattern s9999999999
      ProcessValue <- "86_Times_STEP_MAX_TIME_STP_180(2)"
   AlarmView "Alarm view_1" at 0,777 size 1280x23